   4067: 'Carrier 63 Spacing Fault', class No Acknowledgement, trigger "DB302_HMI_Faults_Carrier63_Faults_2" bit 2
   4068: 'Carrier 63 Duplicate Carrier Number Fault', class No Acknowledgement, trigger "DB302_HMI_Faults_Carrier63_Faults_2" bit 3
   4069: 'Spare_Fault_4069', class No Acknowledgement, trigger "DB302_HMI_Faults_Carrier63_Faults_2" bit 4
   4070: 'Spare_Fault_4070', class No Acknowledgement, trigger "DB302_HMI_Faults_Carrier63_Faults_2" bit 5
   4071: 'Spare_Fault_4071', class No Acknowledgement, trigger "DB302_HMI_Faults_Carrier63_Faults_2" bit 6
   4072: 'Spare_Fault_4072', class No Acknowledgement, trigger "DB302_HMI_Faults_Carrier63_Faults_2" bit 7
   4073: 'Spare_Fault_4073', class No Acknowledgement, trigger "DB302_HMI_Faults_Carrier63_Faults_2" bit 8
   4074: 'Spare_Fault_4074', class No Acknowledgement, trigger "DB302_HMI_Faults_Carrier63_Faults_2" bit 9
   4075: 'Spare_Fault_4075', class No Acknowledgement, trigger "DB302_HMI_Faults_Carrier63_Faults_2" bit 10
   4076: 'Spare_Fault_4076', class No Acknowledgement, trigger "DB302_HMI_Faults_Carrier63_Faults_2" bit 11
   4077: 'Spare_Fault_4077', class No Acknowledgement, trigger "DB302_HMI_Faults_Carrier63_Faults_2" bit 12
   4078: 'Spare_Fault_4078', class No Acknowledgement, trigger "DB302_HMI_Faults_Carrier63_Faults_2" bit 13
   4079: 'Spare_Fault_4079', class No Acknowledgement, trigger "DB302_HMI_Faults_Carrier63_Faults_2" bit 14
   4080: 'Spare_Fault_4080', class No Acknowledgement, trigger "DB302_HMI_Faults_Carrier63_Faults_2" bit 15
   4081: 'Spare_Fault_4081', class No Acknowledgement, trigger "DB302_HMI_Faults_Carrier63_Faults_3" bit 0
   4082: 'Spare_Fault_4082', class No Acknowledgement, trigger "DB302_HMI_Faults_Carrier63_Faults_3" bit 1
   4083: 'Spare_Fault_4083', class No Acknowledgement, trigger "DB302_HMI_Faults_Carrier63_Faults_3" bit 2
   4084: 'Spare_Fault_4084', class No Acknowledgement, trigger "DB302_HMI_Faults_Carrier63_Faults_3" bit 3
   4085: 'Spare_Fault_4085', class No Acknowledgement, trigger "DB302_HMI_Faults_Carrier63_Faults_3" bit 4
   4086: 'Spare_Fault_4086', class No Acknowledgement, trigger "DB302_HMI_Faults_Carrier63_Faults_3" bit 5
   4087: 'Spare_Fault_4087', class No Acknowledgement, trigger "DB302_HMI_Faults_Carrier63_Faults_3" bit 6
   4088: 'Spare_Fault_4088', class No Acknowledgement, trigger "DB302_HMI_Faults_Carrier63_Faults_3" bit 7
   4089: 'Spare_Fault_4089', class No Acknowledgement, trigger "DB302_HMI_Faults_Carrier63_Faults_3" bit 8
   4090: 'Spare_Fault_4090', class No Acknowledgement, trigger "DB302_HMI_Faults_Carrier63_Faults_3" bit 9
   4091: 'Spare_Fault_4091', class No Acknowledgement, trigger "DB302_HMI_Faults_Carrier63_Faults_3" bit 10
   4092: 'Spare_Fault_4092', class No Acknowledgement, trigger "DB302_HMI_Faults_Carrier63_Faults_3" bit 11
   4093: 'Spare_Fault_4093', class No Acknowledgement, trigger "DB302_HMI_Faults_Carrier63_Faults_3" bit 12
   4094: 'Spare_Fault_4094', class No Acknowledgement, trigger "DB302_HMI_Faults_Carrier63_Faults_3" bit 13
   4095: 'Spare_Fault_4095', class No Acknowledgement, trigger "DB302_HMI_Faults_Carrier63_Faults_3" bit 14
   4096: 'Spare_Fault_4096', class No Acknowledgement, trigger "DB302_HMI_Faults_Carrier63_Faults_3" bit 15
   4097: 'Carrier 64 Disconnect Open Power Fault DI11.0', class No Acknowledgement, trigger "DB302_HMI_Faults_Carrier64_Faults_0" bit 0
   4098: 'Carrier 64 Drive Profinet Comm Fault', class No Acknowledgement, trigger "DB302_HMI_Faults_Carrier64_Faults_0" bit 1
   4099: 'Carrier 64 Production Stop Not Reset', class No Acknowledgement, trigger "DB302_HMI_Faults_Carrier64_Faults_0" bit 2
   4100: 'Carrier 64 CB02122 Tripped', class No Acknowledgement, trigger "DB302_HMI_Faults_Carrier64_Faults_0" bit 3
   4101: 'Carrier 64 CB02123 Tripped', class No Acknowledgement, trigger "DB302_HMI_Faults_Carrier64_Faults_0" bit 4
   4102: 'Carrier 64 AUX1 CB Tripped', class No Acknowledgement, trigger "DB302_HMI_Faults_Carrier64_Faults_0" bit 5
   4103: 'Carrier 64 AUX2 CB Tripped', class No Acknowledgement, trigger "DB302_HMI_Faults_Carrier64_Faults_0" bit 6
   4104: 'Carrier 64 PLC Not Communicating', class No Acknowledgement, trigger "DB302_HMI_Faults_Carrier64_Faults_0" bit 7
   4105: 'Carrier 64 Safe Input Card Fault', class No Acknowledgement, trigger "DB302_HMI_Faults_Carrier64_Faults_0" bit 8
   4106: 'Carrier 64 Safe Output Card Fault', class No Acknowledgement, trigger "DB302_HMI_Faults_Carrier64_Faults_0" bit 9
   4107: 'Carrier 64 Standard Input Card Fault', class No Acknowledgement, trigger "DB302_HMI_Faults_Carrier64_Faults_0" bit 10
   4108: 'Carrier 64 Standard Output Card Fault', class No Acknowledgement, trigger "DB302_HMI_Faults_Carrier64_Faults_0" bit 11
   4109: 'Carrier 64 Encoder Position Fault', class No Acknowledgement, trigger "DB302_HMI_Faults_Carrier64_Faults_0" bit 12
   4110: 'Carrier 64 Encoder Internal Error', class No Acknowledgement, trigger "DB302_HMI_Faults_Carrier64_Faults_0" bit 13
   4111: 'Carrier 64 Encoder Comm Fault', class No Acknowledgement, trigger "DB302_HMI_Faults_Carrier64_Faults_0" bit 14
   4112: 'Carrier 64 HMI Comm Fault', class No Acknowledgement, trigger "DB302_HMI_Faults_Carrier64_Faults_0" bit 15
   4113: 'Carrier 64 Crash Detection Fault', class No Acknowledgement, trigger "DB302_HMI_Faults_Carrier64_Faults_1" bit 0
   4114: 'Carrier 64 Carrier Number Invalid', class No Acknowledgement, trigger "DB302_HMI_Faults_Carrier64_Faults_1" bit 1
   4115: 'Carrier 64 Drive: PROFINET configuration error', class No Acknowledgement, trigger "DB302_HMI_Faults_Carrier64_Faults_1" bit 2
   4116: 'Carrier 64 Drive: Error internal communications', class No Acknowledgement, trigger "DB302_HMI_Faults_Carrier64_Faults_1" bit 3
   4117: 'Carrier 64 Drive: Motor overtemperature', class No Acknowledgement, trigger "DB302_HMI_Faults_Carrier64_Faults_1" bit 4
   4118: 'Carrier 64 Drive: Motor overcurrent', class No Acknowledgement, trigger "DB302_HMI_Faults_Carrier64_Faults_1" bit 5
   4119: 'Carrier 64 Drive: Infeed or power unit not ready', class No Acknowledgement, trigger "DB302_HMI_Faults_Carrier64_Faults_1" bit 6
   4120: 'Carrier 64 Drive: Short-circuit/ground fault detected', class No Acknowledgement, trigger "DB302_HMI_Faults_Carrier64_Faults_1" bit 7
   4121: 'Carrier 64 Drive: PROFINET Setpoint timeout', class No Acknowledgement, trigger "DB302_HMI_Faults_Carrier64_Faults_1" bit 8
   4122: 'Carrier 64 Power unit: Overcurrent', class No Acknowledgement, trigger "DB302_HMI_Faults_Carrier64_Faults_1" bit 9
   4123: 'Carrier 64 Power unit: DC link voltage overvoltage', class No Acknowledgement, trigger "DB302_HMI_Faults_Carrier64_Faults_1" bit 10
   4124: 'Carrier 64 Power unit: DC link voltage undervoltage', class No Acknowledgement, trigger "DB302_HMI_Faults_Carrier64_Faults_1" bit 11
   4125: 'Carrier 64 Power unit: Line phase failure in main circuit', class No Acknowledgement, trigger "DB302_HMI_Faults_Carrier64_Faults_1" bit 12
   4126: 'Carrier 64 Power unit: Phase failure motor cable', class No Acknowledgement, trigger "DB302_HMI_Faults_Carrier64_Faults_1" bit 13
   4127: 'Carrier 64 Power unit: Ground fault', class No Acknowledgement, trigger "DB302_HMI_Faults_Carrier64_Faults_1" bit 14
   4128: 'Spare_Fault_4128', class No Acknowledgement, trigger "DB302_HMI_Faults_Carrier64_Faults_1" bit 15
   4129: 'Carrier 64 Motion Off Fault', class No Acknowledgement, trigger "DB302_HMI_Faults_Carrier64_Faults_2" bit 0
   4130: 'Carrier 64 Motion On Fault', class No Acknowledgement, trigger "DB302_HMI_Faults_Carrier64_Faults_2" bit 1
   4131: 'Carrier 64 Spacing Fault', class No Acknowledgement, trigger "DB302_HMI_Faults_Carrier64_Faults_2" bit 2
   4132: 'Carrier 64 Duplicate Carrier Number Fault', class No Acknowledgement, trigger "DB302_HMI_Faults_Carrier64_Faults_2" bit 3
   4133: 'Spare_Fault_4133', class No Acknowledgement, trigger "DB302_HMI_Faults_Carrier64_Faults_2" bit 4
   4134: 'Spare_Fault_4134', class No Acknowledgement, trigger "DB302_HMI_Faults_Carrier64_Faults_2" bit 5
   4135: 'Spare_Fault_4135', class No Acknowledgement, trigger "DB302_HMI_Faults_Carrier64_Faults_2" bit 6
   4136: 'Spare_Fault_4136', class No Acknowledgement, trigger "DB302_HMI_Faults_Carrier64_Faults_2" bit 7
   4137: 'Spare_Fault_4137', class No Acknowledgement, trigger "DB302_HMI_Faults_Carrier64_Faults_2" bit 8
   4138: 'Spare_Fault_4138', class No Acknowledgement, trigger "DB302_HMI_Faults_Carrier64_Faults_2" bit 9
   4139: 'Spare_Fault_4139', class No Acknowledgement, trigger "DB302_HMI_Faults_Carrier64_Faults_2" bit 10
   4140: 'Spare_Fault_4140', class No Acknowledgement, trigger "DB302_HMI_Faults_Carrier64_Faults_2" bit 11
   4141: 'Spare_Fault_4141', class No Acknowledgement, trigger "DB302_HMI_Faults_Carrier64_Faults_2" bit 12
   4142: 'Spare_Fault_4142', class No Acknowledgement, trigger "DB302_HMI_Faults_Carrier64_Faults_2" bit 13
   4143: 'Spare_Fault_4143', class No Acknowledgement, trigger "DB302_HMI_Faults_Carrier64_Faults_2" bit 14
   4144: 'Spare_Fault_4144', class No Acknowledgement, trigger "DB302_HMI_Faults_Carrier64_Faults_2" bit 15
   4145: 'Spare_Fault_4145', class No Acknowledgement, trigger "DB302_HMI_Faults_Carrier64_Faults_3" bit 0
   4146: 'Spare_Fault_4146', class No Acknowledgement, trigger "DB302_HMI_Faults_Carrier64_Faults_3" bit 1
   4147: 'Spare_Fault_4147', class No Acknowledgement, trigger "DB302_HMI_Faults_Carrier64_Faults_3" bit 2
   4148: 'Spare_Fault_4148', class No Acknowledgement, trigger "DB302_HMI_Faults_Carrier64_Faults_3" bit 3
   4149: 'Spare_Fault_4149', class No Acknowledgement, trigger "DB302_HMI_Faults_Carrier64_Faults_3" bit 4
   4150: 'Spare_Fault_4150', class No Acknowledgement, trigger "DB302_HMI_Faults_Carrier64_Faults_3" bit 5
   4151: 'Spare_Fault_4151', class No Acknowledgement, trigger "DB302_HMI_Faults_Carrier64_Faults_3" bit 6
   4152: 'Spare_Fault_4152', class No Acknowledgement, trigger "DB302_HMI_Faults_Carrier64_Faults_3" bit 7
   4153: 'Spare_Fault_4153', class No Acknowledgement, trigger "DB302_HMI_Faults_Carrier64_Faults_3" bit 8
   4154: 'Spare_Fault_4154', class No Acknowledgement, trigger "DB302_HMI_Faults_Carrier64_Faults_3" bit 9
   4155: 'Spare_Fault_4155', class No Acknowledgement, trigger "DB302_HMI_Faults_Carrier64_Faults_3" bit 10
   4156: 'Spare_Fault_4156', class No Acknowledgement, trigger "DB302_HMI_Faults_Carrier64_Faults_3" bit 11
   4157: 'Spare_Fault_4157', class No Acknowledgement, trigger "DB302_HMI_Faults_Carrier64_Faults_3" bit 12
   4158: 'Spare_Fault_4158', class No Acknowledgement, trigger "DB302_HMI_Faults_Carrier64_Faults_3" bit 13
   4159: 'Spare_Fault_4159', class No Acknowledgement, trigger "DB302_HMI_Faults_Carrier64_Faults_3" bit 14
   4160: 'Spare_Fault_4160', class No Acknowledgement, trigger "DB302_HMI_Faults_Carrier64_Faults_3" bit 15
   4161: 'Carrier 65 Disconnect Open Power Fault DI11.0', class No Acknowledgement, trigger "DB302_HMI_Faults_Carrier65_Faults_0" bit 0
   4162: 'Carrier 65 Drive Profinet Comm Fault', class No Acknowledgement, trigger "DB302_HMI_Faults_Carrier65_Faults_0" bit 1
   4163: 'Carrier 65 Production Stop Not Reset', class No Acknowledgement, trigger "DB302_HMI_Faults_Carrier65_Faults_0" bit 2
   4164: 'Carrier 65 CB02122 Tripped', class No Acknowledgement, trigger "DB302_HMI_Faults_Carrier65_Faults_0" bit 3
   4165: 'Carrier 65 CB02123 Tripped', class No Acknowledgement, trigger "DB302_HMI_Faults_Carrier65_Faults_0" bit 4
   4166: 'Carrier 65 AUX1 CB Tripped', class No Acknowledgement, trigger "DB302_HMI_Faults_Carrier65_Faults_0" bit 5
   4167: 'Carrier 65 AUX2 CB Tripped', class No Acknowledgement, trigger "DB302_HMI_Faults_Carrier65_Faults_0" bit 6
   4168: 'Carrier 65 PLC Not Communicating', class No Acknowledgement, trigger "DB302_HMI_Faults_Carrier65_Faults_0" bit 7
   4169: 'Carrier 65 Safe Input Card Fault', class No Acknowledgement, trigger "DB302_HMI_Faults_Carrier65_Faults_0" bit 8
   4170: 'Carrier 65 Safe Output Card Fault', class No Acknowledgement, trigger "DB302_HMI_Faults_Carrier65_Faults_0" bit 9
   4171: 'Carrier 65 Standard Input Card Fault', class No Acknowledgement, trigger "DB302_HMI_Faults_Carrier65_Faults_0" bit 10
   4172: 'Carrier 65 Standard Output Card Fault', class No Acknowledgement, trigger "DB302_HMI_Faults_Carrier65_Faults_0" bit 11
   4173: 'Carrier 65 Encoder Position Fault', class No Acknowledgement, trigger "DB302_HMI_Faults_Carrier65_Faults_0" bit 12
   4174: 'Carrier 65 Encoder Internal Error', class No Acknowledgement, trigger "DB302_HMI_Faults_Carrier65_Faults_0" bit 13
   4175: 'Carrier 65 Encoder Comm Fault', class No Acknowledgement, trigger "DB302_HMI_Faults_Carrier65_Faults_0" bit 14
   4176: 'Carrier 65 HMI Comm Fault', class No Acknowledgement, trigger "DB302_HMI_Faults_Carrier65_Faults_0" bit 15
   4177: 'Carrier 65 Crash Detection Fault', class No Acknowledgement, trigger "DB302_HMI_Faults_Carrier65_Faults_1" bit 0
   4178: 'Carrier 65 Carrier Number Invalid', class No Acknowledgement, trigger "DB302_HMI_Faults_Carrier65_Faults_1" bit 1
   4179: 'Carrier 65 Drive: PROFINET configuration error', class No Acknowledgement, trigger "DB302_HMI_Faults_Carrier65_Faults_1" bit 2
   4180: 'Carrier 65 Drive: Error internal communications', class No Acknowledgement, trigger "DB302_HMI_Faults_Carrier65_Faults_1" bit 3
   4181: 'Carrier 65 Drive: Motor overtemperature', class No Acknowledgement, trigger "DB302_HMI_Faults_Carrier65_Faults_1" bit 4
   4182: 'Carrier 65 Drive: Motor overcurrent', class No Acknowledgement, trigger "DB302_HMI_Faults_Carrier65_Faults_1" bit 5
   4183: 'Carrier 65 Drive: Infeed or power unit not ready', class No Acknowledgement, trigger "DB302_HMI_Faults_Carrier65_Faults_1" bit 6
   4184: 'Carrier 65 Drive: Short-circuit/ground fault detected', class No Acknowledgement, trigger "DB302_HMI_Faults_Carrier65_Faults_1" bit 7
   4185: 'Carrier 65 Drive: PROFINET Setpoint timeout', class No Acknowledgement, trigger "DB302_HMI_Faults_Carrier65_Faults_1" bit 8
   4186: 'Carrier 65 Power unit: Overcurrent', class No Acknowledgement, trigger "DB302_HMI_Faults_Carrier65_Faults_1" bit 9
   4187: 'Carrier 65 Power unit: DC link voltage overvoltage', class No Acknowledgement, trigger "DB302_HMI_Faults_Carrier65_Faults_1" bit 10
   4188: 'Carrier 65 Power unit: DC link voltage undervoltage', class No Acknowledgement, trigger "DB302_HMI_Faults_Carrier65_Faults_1" bit 11
   4189: 'Carrier 65 Power unit: Line phase failure in main circuit', class No Acknowledgement, trigger "DB302_HMI_Faults_Carrier65_Faults_1" bit 12
   4190: 'Carrier 65 Power unit: Phase failure motor cable', class No Acknowledgement, trigger "DB302_HMI_Faults_Carrier65_Faults_1" bit 13
   4191: 'Carrier 65 Power unit: Ground fault', class No Acknowledgement, trigger "DB302_HMI_Faults_Carrier65_Faults_1" bit 14
   4192: 'Spare_Fault_4192', class No Acknowledgement, trigger "DB302_HMI_Faults_Carrier65_Faults_1" bit 15
   4193: 'Carrier 65 Motion Off Fault', class No Acknowledgement, trigger "DB302_HMI_Faults_Carrier65_Faults_2" bit 0
   4194: 'Carrier 65 Motion On Fault', class No Acknowledgement, trigger "DB302_HMI_Faults_Carrier65_Faults_2" bit 1
   4195: 'Carrier 65 Spacing Fault', class No Acknowledgement, trigger "DB302_HMI_Faults_Carrier65_Faults_2" bit 2
   4196: 'Carrier 65 Duplicate Carrier Number Fault', class No Acknowledgement, trigger "DB302_HMI_Faults_Carrier65_Faults_2" bit 3
   4197: 'Spare_Fault_4197', class No Acknowledgement, trigger "DB302_HMI_Faults_Carrier65_Faults_2" bit 4
   4198: 'Spare_Fault_4198', class No Acknowledgement, trigger "DB302_HMI_Faults_Carrier65_Faults_2" bit 5
   4199: 'Spare_Fault_4199', class No Acknowledgement, trigger "DB302_HMI_Faults_Carrier65_Faults_2" bit 6
   4200: 'Spare_Fault_4200', class No Acknowledgement, trigger "DB302_HMI_Faults_Carrier65_Faults_2" bit 7
   4201: 'Spare_Fault_4201', class No Acknowledgement, trigger "DB302_HMI_Faults_Carrier65_Faults_2" bit 8
   4202: 'Spare_Fault_4202', class No Acknowledgement, trigger "DB302_HMI_Faults_Carrier65_Faults_2" bit 9
   4203: 'Spare_Fault_4203', class No Acknowledgement, trigger "DB302_HMI_Faults_Carrier65_Faults_2" bit 10
   4204: 'Spare_Fault_4204', class No Acknowledgement, trigger "DB302_HMI_Faults_Carrier65_Faults_2" bit 11
   4205: 'Spare_Fault_4205', class No Acknowledgement, trigger "DB302_HMI_Faults_Carrier65_Faults_2" bit 12
   4206: 'Spare_Fault_4206', class No Acknowledgement, trigger "DB302_HMI_Faults_Carrier65_Faults_2" bit 13
   4207: 'Spare_Fault_4207', class No Acknowledgement, trigger "DB302_HMI_Faults_Carrier65_Faults_2" bit 14
   4208: 'Spare_Fault_4208', class No Acknowledgement, trigger "DB302_HMI_Faults_Carrier65_Faults_2" bit 15
   4209: 'Spare_Fault_4209', class No Acknowledgement, trigger "DB302_HMI_Faults_Carrier65_Faults_3" bit 0
   4210: 'Spare_Fault_4210', class No Acknowledgement, trigger "DB302_HMI_Faults_Carrier65_Faults_3" bit 1
   4211: 'Spare_Fault_4211', class No Acknowledgement, trigger "DB302_HMI_Faults_Carrier65_Faults_3" bit 2
   4212: 'Spare_Fault_4212', class No Acknowledgement, trigger "DB302_HMI_Faults_Carrier65_Faults_3" bit 3
   4213: 'Spare_Fault_4213', class No Acknowledgement, trigger "DB302_HMI_Faults_Carrier65_Faults_3" bit 4
   4214: 'Spare_Fault_4214', class No Acknowledgement, trigger "DB302_HMI_Faults_Carrier65_Faults_3" bit 5
   4215: 'Spare_Fault_4215', class No Acknowledgement, trigger "DB302_HMI_Faults_Carrier65_Faults_3" bit 6
   4216: 'Spare_Fault_4216', class No Acknowledgement, trigger "DB302_HMI_Faults_Carrier65_Faults_3" bit 7
   4217: 'Spare_Fault_4217', class No Acknowledgement, trigger "DB302_HMI_Faults_Carrier65_Faults_3" bit 8
   4218: 'Spare_Fault_4218', class No Acknowledgement, trigger "DB302_HMI_Faults_Carrier65_Faults_3" bit 9
   4219: 'Spare_Fault_4219', class No Acknowledgement, trigger "DB302_HMI_Faults_Carrier65_Faults_3" bit 10
   4220: 'Spare_Fault_4220', class No Acknowledgement, trigger "DB302_HMI_Faults_Carrier65_Faults_3" bit 11
   4221: 'Spare_Fault_4221', class No Acknowledgement, trigger "DB302_HMI_Faults_Carrier65_Faults_3" bit 12
   4222: 'Spare_Fault_4222', class No Acknowledgement, trigger "DB302_HMI_Faults_Carrier65_Faults_3" bit 13
   4223: 'Spare_Fault_4223', class No Acknowledgement, trigger "DB302_HMI_Faults_Carrier65_Faults_3" bit 14
   4224: 'Spare_Fault_4224', class No Acknowledgement, trigger "DB302_HMI_Faults_Carrier65_Faults_3" bit 15
   4225: 'Carrier 66 Disconnect Open Power Fault DI11.0', class No Acknowledgement, trigger "DB302_HMI_Faults_Carrier66_Faults_0" bit 0
   4226: 'Carrier 66 Drive Profinet Comm Fault', class No Acknowledgement, trigger "DB302_HMI_Faults_Carrier66_Faults_0" bit 1
   4227: 'Carrier 66 Production Stop Not Reset', class No Acknowledgement, trigger "DB302_HMI_Faults_Carrier66_Faults_0" bit 2
   4228: 'Carrier 66 CB02122 Tripped', class No Acknowledgement, trigger "DB302_HMI_Faults_Carrier66_Faults_0" bit 3
   4229: 'Carrier 66 CB02123 Tripped', class No Acknowledgement, trigger "DB302_HMI_Faults_Carrier66_Faults_0" bit 4
   4230: 'Carrier 66 AUX1 CB Tripped', class No Acknowledgement, trigger "DB302_HMI_Faults_Carrier66_Faults_0" bit 5
   4231: 'Carrier 66 AUX2 CB Tripped', class No Acknowledgement, trigger "DB302_HMI_Faults_Carrier66_Faults_0" bit 6
   4232: 'Carrier 66 PLC Not Communicating', class No Acknowledgement, trigger "DB302_HMI_Faults_Carrier66_Faults_0" bit 7
   4233: 'Carrier 66 Safe Input Card Fault', class No Acknowledgement, trigger "DB302_HMI_Faults_Carrier66_Faults_0" bit 8
   4234: 'Carrier 66 Safe Output Card Fault', class No Acknowledgement, trigger "DB302_HMI_Faults_Carrier66_Faults_0" bit 9
   4235: 'Carrier 66 Standard Input Card Fault', class No Acknowledgement, trigger "DB302_HMI_Faults_Carrier66_Faults_0" bit 10
   4236: 'Carrier 66 Standard Output Card Fault', class No Acknowledgement, trigger "DB302_HMI_Faults_Carrier66_Faults_0" bit 11
   4237: 'Carrier 66 Encoder Position Fault', class No Acknowledgement, trigger "DB302_HMI_Faults_Carrier66_Faults_0" bit 12
   4238: 'Carrier 66 Encoder Internal Error', class No Acknowledgement, trigger "DB302_HMI_Faults_Carrier66_Faults_0" bit 13
   4239: 'Carrier 66 Encoder Comm Fault', class No Acknowledgement, trigger "DB302_HMI_Faults_Carrier66_Faults_0" bit 14
   4240: 'Carrier 66 HMI Comm Fault', class No Acknowledgement, trigger "DB302_HMI_Faults_Carrier66_Faults_0" bit 15
   4241: 'Carrier 66 Crash Detection Fault', class No Acknowledgement, trigger "DB302_HMI_Faults_Carrier66_Faults_1" bit 0
   4242: 'Carrier 66 Carrier Number Invalid', class No Acknowledgement, trigger "DB302_HMI_Faults_Carrier66_Faults_1" bit 1
   4243: 'Carrier 66 Drive: PROFINET configuration error', class No Acknowledgement, trigger "DB302_HMI_Faults_Carrier66_Faults_1" bit 2
   4244: 'Carrier 66 Drive: Error internal communications', class No Acknowledgement, trigger "DB302_HMI_Faults_Carrier66_Faults_1" bit 3
   4245: 'Carrier 66 Drive: Motor overtemperature', class No Acknowledgement, trigger "DB302_HMI_Faults_Carrier66_Faults_1" bit 4
   4246: 'Carrier 66 Drive: Motor overcurrent', class No Acknowledgement, trigger "DB302_HMI_Faults_Carrier66_Faults_1" bit 5
   4247: 'Carrier 66 Drive: Infeed or power unit not ready', class No Acknowledgement, trigger "DB302_HMI_Faults_Carrier66_Faults_1" bit 6
   4248: 'Carrier 66 Drive: Short-circuit/ground fault detected', class No Acknowledgement, trigger "DB302_HMI_Faults_Carrier66_Faults_1" bit 7
   4249: 'Carrier 66 Drive: PROFINET Setpoint timeout', class No Acknowledgement, trigger "DB302_HMI_Faults_Carrier66_Faults_1" bit 8
   4250: 'Carrier 66 Power unit: Overcurrent', class No Acknowledgement, trigger "DB302_HMI_Faults_Carrier66_Faults_1" bit 9
   4251: 'Carrier 66 Power unit: DC link voltage overvoltage', class No Acknowledgement, trigger "DB302_HMI_Faults_Carrier66_Faults_1" bit 10
   4252: 'Carrier 66 Power unit: DC link voltage undervoltage', class No Acknowledgement, trigger "DB302_HMI_Faults_Carrier66_Faults_1" bit 11
   4253: 'Carrier 66 Power unit: Line phase failure in main circuit', class No Acknowledgement, trigger "DB302_HMI_Faults_Carrier66_Faults_1" bit 12
   4254: 'Carrier 66 Power unit: Phase failure motor cable', class No Acknowledgement, trigger "DB302_HMI_Faults_Carrier66_Faults_1" bit 13
   4255: 'Carrier 66 Power unit: Ground fault', class No Acknowledgement, trigger "DB302_HMI_Faults_Carrier66_Faults_1" bit 14
   4256: 'Spare_Fault_4256', class No Acknowledgement, trigger "DB302_HMI_Faults_Carrier66_Faults_1" bit 15
   4257: 'Carrier 66 Motion Off Fault', class No Acknowledgement, trigger "DB302_HMI_Faults_Carrier66_Faults_2" bit 0
   4258: 'Carrier 66 Motion On Fault', class No Acknowledgement, trigger "DB302_HMI_Faults_Carrier66_Faults_2" bit 1
   4259: 'Carrier 66 Spacing Fault', class No Acknowledgement, trigger "DB302_HMI_Faults_Carrier66_Faults_2" bit 2
   4260: 'Carrier 66 Duplicate Carrier Number Fault', class No Acknowledgement, trigger "DB302_HMI_Faults_Carrier66_Faults_2" bit 3
   4261: 'Spare_Fault_4261', class No Acknowledgement, trigger "DB302_HMI_Faults_Carrier66_Faults_2" bit 4
   4262: 'Spare_Fault_4262', class No Acknowledgement, trigger "DB302_HMI_Faults_Carrier66_Faults_2" bit 5
   4263: 'Spare_Fault_4263', class No Acknowledgement, trigger "DB302_HMI_Faults_Carrier66_Faults_2" bit 6
   4264: 'Spare_Fault_4264', class No Acknowledgement, trigger "DB302_HMI_Faults_Carrier66_Faults_2" bit 7
   4265: 'Spare_Fault_4265', class No Acknowledgement, trigger "DB302_HMI_Faults_Carrier66_Faults_2" bit 8
   4266: 'Spare_Fault_4266', class No Acknowledgement, trigger "DB302_HMI_Faults_Carrier66_Faults_2" bit 9
   4267: 'Spare_Fault_4267', class No Acknowledgement, trigger "DB302_HMI_Faults_Carrier66_Faults_2" bit 10
   4268: 'Spare_Fault_4268', class No Acknowledgement, trigger "DB302_HMI_Faults_Carrier66_Faults_2" bit 11
   4269: 'Spare_Fault_4269', class No Acknowledgement, trigger "DB302_HMI_Faults_Carrier66_Faults_2" bit 12
   4270: 'Spare_Fault_4270', class No Acknowledgement, trigger "DB302_HMI_Faults_Carrier66_Faults_2" bit 13
   4271: 'Spare_Fault_4271', class No Acknowledgement, trigger "DB302_HMI_Faults_Carrier66_Faults_2" bit 14
   4272: 'Spare_Fault_4272', class No Acknowledgement, trigger "DB302_HMI_Faults_Carrier66_Faults_2" bit 15
   4273: 'Spare_Fault_4273', class No Acknowledgement, trigger "DB302_HMI_Faults_Carrier66_Faults_3" bit 0
   4274: 'Spare_Fault_4274', class No Acknowledgement, trigger "DB302_HMI_Faults_Carrier66_Faults_3" bit 1
   4275: 'Spare_Fault_4275', class No Acknowledgement, trigger "DB302_HMI_Faults_Carrier66_Faults_3" bit 2
   4276: 'Spare_Fault_4276', class No Acknowledgement, trigger "DB302_HMI_Faults_Carrier66_Faults_3" bit 3
   4277: 'Spare_Fault_4277', class No Acknowledgement, trigger "DB302_HMI_Faults_Carrier66_Faults_3" bit 4
   4278: 'Spare_Fault_4278', class No Acknowledgement, trigger "DB302_HMI_Faults_Carrier66_Faults_3" bit 5
   4279: 'Spare_Fault_4279', class No Acknowledgement, trigger "DB302_HMI_Faults_Carrier66_Faults_3" bit 6
   4280: 'Spare_Fault_4280', class No Acknowledgement, trigger "DB302_HMI_Faults_Carrier66_Faults_3" bit 7
   4281: 'Spare_Fault_4281', class No Acknowledgement, trigger "DB302_HMI_Faults_Carrier66_Faults_3" bit 8
   4282: 'Spare_Fault_4282', class No Acknowledgement, trigger "DB302_HMI_Faults_Carrier66_Faults_3" bit 9
   4283: 'Spare_Fault_4283', class No Acknowledgement, trigger "DB302_HMI_Faults_Carrier66_Faults_3" bit 10
   4284: 'Spare_Fault_4284', class No Acknowledgement, trigger "DB302_HMI_Faults_Carrier66_Faults_3" bit 11
   4285: 'Spare_Fault_4285', class No Acknowledgement, trigger "DB302_HMI_Faults_Carrier66_Faults_3" bit 12
   4286: 'Spare_Fault_4286', class No Acknowledgement, trigger "DB302_HMI_Faults_Carrier66_Faults_3" bit 13
   4287: 'Spare_Fault_4287', class No Acknowledgement, trigger "DB302_HMI_Faults_Carrier66_Faults_3" bit 14
   4288: 'Spare_Fault_4288', class No Acknowledgement, trigger "DB302_HMI_Faults_Carrier66_Faults_3" bit 15
   4289: 'Carrier 67 Disconnect Open Power Fault DI11.0', class No Acknowledgement, trigger "DB302_HMI_Faults_Carrier67_Faults_0" bit 0
   4290: 'Carrier 67 Drive Profinet Comm Fault', class No Acknowledgement, trigger "DB302_HMI_Faults_Carrier67_Faults_0" bit 1
   4291: 'Carrier 67 Production Stop Not Reset', class No Acknowledgement, trigger "DB302_HMI_Faults_Carrier67_Faults_0" bit 2
   4292: 'Carrier 67 CB02122 Tripped', class No Acknowledgement, trigger "DB302_HMI_Faults_Carrier67_Faults_0" bit 3
   4293: 'Carrier 67 CB02123 Tripped', class No Acknowledgement, trigger "DB302_HMI_Faults_Carrier67_Faults_0" bit 4
   4294: 'Carrier 67 AUX1 CB Tripped', class No Acknowledgement, trigger "DB302_HMI_Faults_Carrier67_Faults_0" bit 5
   4295: 'Carrier 67 AUX2 CB Tripped', class No Acknowledgement, trigger "DB302_HMI_Faults_Carrier67_Faults_0" bit 6
   4296: 'Carrier 67 PLC Not Communicating', class No Acknowledgement, trigger "DB302_HMI_Faults_Carrier67_Faults_0" bit 7
   4297: 'Carrier 67 Safe Input Card Fault', class No Acknowledgement, trigger "DB302_HMI_Faults_Carrier67_Faults_0" bit 8
   4298: 'Carrier 67 Safe Output Card Fault', class No Acknowledgement, trigger "DB302_HMI_Faults_Carrier67_Faults_0" bit 9
   4299: 'Carrier 67 Standard Input Card Fault', class No Acknowledgement, trigger "DB302_HMI_Faults_Carrier67_Faults_0" bit 10
   4300: 'Carrier 67 Standard Output Card Fault', class No Acknowledgement, trigger "DB302_HMI_Faults_Carrier67_Faults_0" bit 11
   4301: 'Carrier 67 Encoder Position Fault', class No Acknowledgement, trigger "DB302_HMI_Faults_Carrier67_Faults_0" bit 12
   4302: 'Carrier 67 Encoder Internal Error', class No Acknowledgement, trigger "DB302_HMI_Faults_Carrier67_Faults_0" bit 13
   4303: 'Carrier 67 Encoder Comm Fault', class No Acknowledgement, trigger "DB302_HMI_Faults_Carrier67_Faults_0" bit 14
   4304: 'Carrier 67 HMI Comm Fault', class No Acknowledgement, trigger "DB302_HMI_Faults_Carrier67_Faults_0" bit 15
   4305: 'Carrier 67 Crash Detection Fault', class No Acknowledgement, trigger "DB302_HMI_Faults_Carrier67_Faults_1" bit 0
   4306: 'Carrier 67 Carrier Number Invalid', class No Acknowledgement, trigger "DB302_HMI_Faults_Carrier67_Faults_1" bit 1
   4307: 'Carrier 67 Drive: PROFINET configuration error', class No Acknowledgement, trigger "DB302_HMI_Faults_Carrier67_Faults_1" bit 2
   4308: 'Carrier 67 Drive: Error internal communications', class No Acknowledgement, trigger "DB302_HMI_Faults_Carrier67_Faults_1" bit 3
   4309: 'Carrier 67 Drive: Motor overtemperature', class No Acknowledgement, trigger "DB302_HMI_Faults_Carrier67_Faults_1" bit 4
   4310: 'Carrier 67 Drive: Motor overcurrent', class No Acknowledgement, trigger "DB302_HMI_Faults_Carrier67_Faults_1" bit 5
   4311: 'Carrier 67 Drive: Infeed or power unit not ready', class No Acknowledgement, trigger "DB302_HMI_Faults_Carrier67_Faults_1" bit 6
   4312: 'Carrier 67 Drive: Short-circuit/ground fault detected', class No Acknowledgement, trigger "DB302_HMI_Faults_Carrier67_Faults_1" bit 7
   4313: 'Carrier 67 Drive: PROFINET Setpoint timeout', class No Acknowledgement, trigger "DB302_HMI_Faults_Carrier67_Faults_1" bit 8
   4314: 'Carrier 67 Power unit: Overcurrent', class No Acknowledgement, trigger "DB302_HMI_Faults_Carrier67_Faults_1" bit 9
   4315: 'Carrier 67 Power unit: DC link voltage overvoltage', class No Acknowledgement, trigger "DB302_HMI_Faults_Carrier67_Faults_1" bit 10
   4316: 'Carrier 67 Power unit: DC link voltage undervoltage', class No Acknowledgement, trigger "DB302_HMI_Faults_Carrier67_Faults_1" bit 11
   4317: 'Carrier 67 Power unit: Line phase failure in main circuit', class No Acknowledgement, trigger "DB302_HMI_Faults_Carrier67_Faults_1" bit 12
   4318: 'Carrier 67 Power unit: Phase failure motor cable', class No Acknowledgement, trigger "DB302_HMI_Faults_Carrier67_Faults_1" bit 13
   4319: 'Carrier 67 Power unit: Ground fault', class No Acknowledgement, trigger "DB302_HMI_Faults_Carrier67_Faults_1" bit 14
   4320: 'Spare_Fault_4320', class No Acknowledgement, trigger "DB302_HMI_Faults_Carrier67_Faults_1" bit 15
   4321: 'Carrier 67 Motion Off Fault', class No Acknowledgement, trigger "DB302_HMI_Faults_Carrier67_Faults_2" bit 0
   4322: 'Carrier 67 Motion On Fault', class No Acknowledgement, trigger "DB302_HMI_Faults_Carrier67_Faults_2" bit 1
   4323: 'Carrier 67 Spacing Fault', class No Acknowledgement, trigger "DB302_HMI_Faults_Carrier67_Faults_2" bit 2
   4324: 'Carrier 67 Duplicate Carrier Number Fault', class No Acknowledgement, trigger "DB302_HMI_Faults_Carrier67_Faults_2" bit 3
   4325: 'Spare_Fault_4325', class No Acknowledgement, trigger "DB302_HMI_Faults_Carrier67_Faults_2" bit 4
   4326: 'Spare_Fault_4326', class No Acknowledgement, trigger "DB302_HMI_Faults_Carrier67_Faults_2" bit 5
   4327: 'Spare_Fault_4327', class No Acknowledgement, trigger "DB302_HMI_Faults_Carrier67_Faults_2" bit 6
   4328: 'Spare_Fault_4328', class No Acknowledgement, trigger "DB302_HMI_Faults_Carrier67_Faults_2" bit 7
   4329: 'Spare_Fault_4329', class No Acknowledgement, trigger "DB302_HMI_Faults_Carrier67_Faults_2" bit 8
   4330: 'Spare_Fault_4330', class No Acknowledgement, trigger "DB302_HMI_Faults_Carrier67_Faults_2" bit 9
   4331: 'Spare_Fault_4331', class No Acknowledgement, trigger "DB302_HMI_Faults_Carrier67_Faults_2" bit 10
   4332: 'Spare_Fault_4332', class No Acknowledgement, trigger "DB302_HMI_Faults_Carrier67_Faults_2" bit 11
   4333: 'Spare_Fault_4333', class No Acknowledgement, trigger "DB302_HMI_Faults_Carrier67_Faults_2" bit 12
   4334: 'Spare_Fault_4334', class No Acknowledgement, trigger "DB302_HMI_Faults_Carrier67_Faults_2" bit 13
   4335: 'Spare_Fault_4335', class No Acknowledgement, trigger "DB302_HMI_Faults_Carrier67_Faults_2" bit 14
   4336: 'Spare_Fault_4336', class No Acknowledgement, trigger "DB302_HMI_Faults_Carrier67_Faults_2" bit 15
   4337: 'Spare_Fault_4337', class No Acknowledgement, trigger "DB302_HMI_Faults_Carrier67_Faults_3" bit 0
   4338: 'Spare_Fault_4338', class No Acknowledgement, trigger "DB302_HMI_Faults_Carrier67_Faults_3" bit 1
   4339: 'Spare_Fault_4339', class No Acknowledgement, trigger "DB302_HMI_Faults_Carrier67_Faults_3" bit 2
   4340: 'Spare_Fault_4340', class No Acknowledgement, trigger "DB302_HMI_Faults_Carrier67_Faults_3" bit 3
   4341: 'Spare_Fault_4341', class No Acknowledgement, trigger "DB302_HMI_Faults_Carrier67_Faults_3" bit 4
   4342: 'Spare_Fault_4342', class No Acknowledgement, trigger "DB302_HMI_Faults_Carrier67_Faults_3" bit 5
   4343: 'Spare_Fault_4343', class No Acknowledgement, trigger "DB302_HMI_Faults_Carrier67_Faults_3" bit 6
   4344: 'Spare_Fault_4344', class No Acknowledgement, trigger "DB302_HMI_Faults_Carrier67_Faults_3" bit 7
   4345: 'Spare_Fault_4345', class No Acknowledgement, trigger "DB302_HMI_Faults_Carrier67_Faults_3" bit 8
   4346: 'Spare_Fault_4346', class No Acknowledgement, trigger "DB302_HMI_Faults_Carrier67_Faults_3" bit 9
   4347: 'Spare_Fault_4347', class No Acknowledgement, trigger "DB302_HMI_Faults_Carrier67_Faults_3" bit 10
   4348: 'Spare_Fault_4348', class No Acknowledgement, trigger "DB302_HMI_Faults_Carrier67_Faults_3" bit 11
   4349: 'Spare_Fault_4349', class No Acknowledgement, trigger "DB302_HMI_Faults_Carrier67_Faults_3" bit 12
   4350: 'Spare_Fault_4350', class No Acknowledgement, trigger "DB302_HMI_Faults_Carrier67_Faults_3" bit 13
   4351: 'Spare_Fault_4351', class No Acknowledgement, trigger "DB302_HMI_Faults_Carrier67_Faults_3" bit 14
   4352: 'Spare_Fault_4352', class No Acknowledgement, trigger "DB302_HMI_Faults_Carrier67_Faults_3" bit 15
   4353: 'Carrier 68 Disconnect Open Power Fault DI11.0', class No Acknowledgement, trigger "DB302_HMI_Faults_Carrier68_Faults_0" bit 0
   4354: 'Carrier 68 Drive Profinet Comm Fault', class No Acknowledgement, trigger "DB302_HMI_Faults_Carrier68_Faults_0" bit 1
   4355: 'Carrier 68 Production Stop Not Reset', class No Acknowledgement, trigger "DB302_HMI_Faults_Carrier68_Faults_0" bit 2
   4356: 'Carrier 68 CB02122 Tripped', class No Acknowledgement, trigger "DB302_HMI_Faults_Carrier68_Faults_0" bit 3
   4357: 'Carrier 68 CB02123 Tripped', class No Acknowledgement, trigger "DB302_HMI_Faults_Carrier68_Faults_0" bit 4
   4358: 'Carrier 68 AUX1 CB Tripped', class No Acknowledgement, trigger "DB302_HMI_Faults_Carrier68_Faults_0" bit 5
   4359: 'Carrier 68 AUX2 CB Tripped', class No Acknowledgement, trigger "DB302_HMI_Faults_Carrier68_Faults_0" bit 6
   4360: 'Carrier 68 PLC Not Communicating', class No Acknowledgement, trigger "DB302_HMI_Faults_Carrier68_Faults_0" bit 7
   4361: 'Carrier 68 Safe Input Card Fault', class No Acknowledgement, trigger "DB302_HMI_Faults_Carrier68_Faults_0" bit 8
   4362: 'Carrier 68 Safe Output Card Fault', class No Acknowledgement, trigger "DB302_HMI_Faults_Carrier68_Faults_0" bit 9
   4363: 'Carrier 68 Standard Input Card Fault', class No Acknowledgement, trigger "DB302_HMI_Faults_Carrier68_Faults_0" bit 10
   4364: 'Carrier 68 Standard Output Card Fault', class No Acknowledgement, trigger "DB302_HMI_Faults_Carrier68_Faults_0" bit 11
   4365: 'Carrier 68 Encoder Position Fault', class No Acknowledgement, trigger "DB302_HMI_Faults_Carrier68_Faults_0" bit 12
   4366: 'Carrier 68 Encoder Internal Error', class No Acknowledgement, trigger "DB302_HMI_Faults_Carrier68_Faults_0" bit 13
   4367: 'Carrier 68 Encoder Comm Fault', class No Acknowledgement, trigger "DB302_HMI_Faults_Carrier68_Faults_0" bit 14
   4368: 'Carrier 68 HMI Comm Fault', class No Acknowledgement, trigger "DB302_HMI_Faults_Carrier68_Faults_0" bit 15
   4369: 'Carrier 68 Crash Detection Fault', class No Acknowledgement, trigger "DB302_HMI_Faults_Carrier68_Faults_1" bit 0
   4370: 'Carrier 68 Carrier Number Invalid', class No Acknowledgement, trigger "DB302_HMI_Faults_Carrier68_Faults_1" bit 1
   4371: 'Carrier 68 Drive: PROFINET configuration error', class No Acknowledgement, trigger "DB302_HMI_Faults_Carrier68_Faults_1" bit 2
   4372: 'Carrier 68 Drive: Error internal communications', class No Acknowledgement, trigger "DB302_HMI_Faults_Carrier68_Faults_1" bit 3
   4373: 'Carrier 68 Drive: Motor overtemperature', class No Acknowledgement, trigger "DB302_HMI_Faults_Carrier68_Faults_1" bit 4
   4374: 'Carrier 68 Drive: Motor overcurrent', class No Acknowledgement, trigger "DB302_HMI_Faults_Carrier68_Faults_1" bit 5
   4375: 'Carrier 68 Drive: Infeed or power unit not ready', class No Acknowledgement, trigger "DB302_HMI_Faults_Carrier68_Faults_1" bit 6
   4376: 'Carrier 68 Drive: Short-circuit/ground fault detected', class No Acknowledgement, trigger "DB302_HMI_Faults_Carrier68_Faults_1" bit 7
   4377: 'Carrier 68 Drive: PROFINET Setpoint timeout', class No Acknowledgement, trigger "DB302_HMI_Faults_Carrier68_Faults_1" bit 8
   4378: 'Carrier 68 Power unit: Overcurrent', class No Acknowledgement, trigger "DB302_HMI_Faults_Carrier68_Faults_1" bit 9
   4379: 'Carrier 68 Power unit: DC link voltage overvoltage', class No Acknowledgement, trigger "DB302_HMI_Faults_Carrier68_Faults_1" bit 10
   4380: 'Carrier 68 Power unit: DC link voltage undervoltage', class No Acknowledgement, trigger "DB302_HMI_Faults_Carrier68_Faults_1" bit 11
   4381: 'Carrier 68 Power unit: Line phase failure in main circuit', class No Acknowledgement, trigger "DB302_HMI_Faults_Carrier68_Faults_1" bit 12
   4382: 'Carrier 68 Power unit: Phase failure motor cable', class No Acknowledgement, trigger "DB302_HMI_Faults_Carrier68_Faults_1" bit 13
   4383: 'Carrier 68 Power unit: Ground fault', class No Acknowledgement, trigger "DB302_HMI_Faults_Carrier68_Faults_1" bit 14
   4384: 'Spare_Fault_4384', class No Acknowledgement, trigger "DB302_HMI_Faults_Carrier68_Faults_1" bit 15
   4385: 'Carrier 68 Motion Off Fault', class No Acknowledgement, trigger "DB302_HMI_Faults_Carrier68_Faults_2" bit 0
   4386: 'Carrier 68 Motion On Fault', class No Acknowledgement, trigger "DB302_HMI_Faults_Carrier68_Faults_2" bit 1
   4387: 'Carrier 68 Spacing Fault', class No Acknowledgement, trigger "DB302_HMI_Faults_Carrier68_Faults_2" bit 2
   4388: 'Carrier 68 Duplicate Carrier Number Fault', class No Acknowledgement, trigger "DB302_HMI_Faults_Carrier68_Faults_2" bit 3
   4389: 'Spare_Fault_4389', class No Acknowledgement, trigger "DB302_HMI_Faults_Carrier68_Faults_2" bit 4
   4390: 'Spare_Fault_4390', class No Acknowledgement, trigger "DB302_HMI_Faults_Carrier68_Faults_2" bit 5
   4391: 'Spare_Fault_4391', class No Acknowledgement, trigger "DB302_HMI_Faults_Carrier68_Faults_2" bit 6
   4392: 'Spare_Fault_4392', class No Acknowledgement, trigger "DB302_HMI_Faults_Carrier68_Faults_2" bit 7
   4393: 'Spare_Fault_4393', class No Acknowledgement, trigger "DB302_HMI_Faults_Carrier68_Faults_2" bit 8
   4394: 'Spare_Fault_4394', class No Acknowledgement, trigger "DB302_HMI_Faults_Carrier68_Faults_2" bit 9
   4395: 'Spare_Fault_4395', class No Acknowledgement, trigger "DB302_HMI_Faults_Carrier68_Faults_2" bit 10
   4396: 'Spare_Fault_4396', class No Acknowledgement, trigger "DB302_HMI_Faults_Carrier68_Faults_2" bit 11
   4397: 'Spare_Fault_4397', class No Acknowledgement, trigger "DB302_HMI_Faults_Carrier68_Faults_2" bit 12
   4398: 'Spare_Fault_4398', class No Acknowledgement, trigger "DB302_HMI_Faults_Carrier68_Faults_2" bit 13
   4399: 'Spare_Fault_4399', class No Acknowledgement, trigger "DB302_HMI_Faults_Carrier68_Faults_2" bit 14
   4400: 'Spare_Fault_4400', class No Acknowledgement, trigger "DB302_HMI_Faults_Carrier68_Faults_2" bit 15
   4401: 'Spare_Fault_4401', class No Acknowledgement, trigger "DB302_HMI_Faults_Carrier68_Faults_3" bit 0
   4402: 'Spare_Fault_4402', class No Acknowledgement, trigger "DB302_HMI_Faults_Carrier68_Faults_3" bit 1
   4403: 'Spare_Fault_4403', class No Acknowledgement, trigger "DB302_HMI_Faults_Carrier68_Faults_3" bit 2
   4404: 'Spare_Fault_4404', class No Acknowledgement, trigger "DB302_HMI_Faults_Carrier68_Faults_3" bit 3
   4405: 'Spare_Fault_4405', class No Acknowledgement, trigger "DB302_HMI_Faults_Carrier68_Faults_3" bit 4
   4406: 'Spare_Fault_4406', class No Acknowledgement, trigger "DB302_HMI_Faults_Carrier68_Faults_3" bit 5
   4407: 'Spare_Fault_4407', class No Acknowledgement, trigger "DB302_HMI_Faults_Carrier68_Faults_3" bit 6
   4408: 'Spare_Fault_4408', class No Acknowledgement, trigger "DB302_HMI_Faults_Carrier68_Faults_3" bit 7
   4409: 'Spare_Fault_4409', class No Acknowledgement, trigger "DB302_HMI_Faults_Carrier68_Faults_3" bit 8
   4410: 'Spare_Fault_4410', class No Acknowledgement, trigger "DB302_HMI_Faults_Carrier68_Faults_3" bit 9
   4411: 'Spare_Fault_4411', class No Acknowledgement, trigger "DB302_HMI_Faults_Carrier68_Faults_3" bit 10
   4412: 'Spare_Fault_4412', class No Acknowledgement, trigger "DB302_HMI_Faults_Carrier68_Faults_3" bit 11
   4413: 'Spare_Fault_4413', class No Acknowledgement, trigger "DB302_HMI_Faults_Carrier68_Faults_3" bit 12
   4414: 'Spare_Fault_4414', class No Acknowledgement, trigger "DB302_HMI_Faults_Carrier68_Faults_3" bit 13
   4415: 'Spare_Fault_4415', class No Acknowledgement, trigger "DB302_HMI_Faults_Carrier68_Faults_3" bit 14
   4416: 'Spare_Fault_4416', class No Acknowledgement, trigger "DB302_HMI_Faults_Carrier68_Faults_3" bit 15
   4417: 'Carrier 69 Disconnect Open Power Fault DI11.0', class No Acknowledgement, trigger "DB302_HMI_Faults_Carrier69_Faults_0" bit 0
   4418: 'Carrier 69 Drive Profinet Comm Fault', class No Acknowledgement, trigger "DB302_HMI_Faults_Carrier69_Faults_0" bit 1
   4419: 'Carrier 69 Production Stop Not Reset', class No Acknowledgement, trigger "DB302_HMI_Faults_Carrier69_Faults_0" bit 2
   4420: 'Carrier 69 CB02122 Tripped', class No Acknowledgement, trigger "DB302_HMI_Faults_Carrier69_Faults_0" bit 3
   4421: 'Carrier 69 CB02123 Tripped', class No Acknowledgement, trigger "DB302_HMI_Faults_Carrier69_Faults_0" bit 4
   4422: 'Carrier 69 AUX1 CB Tripped', class No Acknowledgement, trigger "DB302_HMI_Faults_Carrier69_Faults_0" bit 5
   4423: 'Carrier 69 AUX2 CB Tripped', class No Acknowledgement, trigger "DB302_HMI_Faults_Carrier69_Faults_0" bit 6
   4424: 'Carrier 69 PLC Not Communicating', class No Acknowledgement, trigger "DB302_HMI_Faults_Carrier69_Faults_0" bit 7
   4425: 'Carrier 69 Safe Input Card Fault', class No Acknowledgement, trigger "DB302_HMI_Faults_Carrier69_Faults_0" bit 8
   4426: 'Carrier 69 Safe Output Card Fault', class No Acknowledgement, trigger "DB302_HMI_Faults_Carrier69_Faults_0" bit 9
   4427: 'Carrier 69 Standard Input Card Fault', class No Acknowledgement, trigger "DB302_HMI_Faults_Carrier69_Faults_0" bit 10
   4428: 'Carrier 69 Standard Output Card Fault', class No Acknowledgement, trigger "DB302_HMI_Faults_Carrier69_Faults_0" bit 11
   4429: 'Carrier 69 Encoder Position Fault', class No Acknowledgement, trigger "DB302_HMI_Faults_Carrier69_Faults_0" bit 12
   4430: 'Carrier 69 Encoder Internal Error', class No Acknowledgement, trigger "DB302_HMI_Faults_Carrier69_Faults_0" bit 13
   4431: 'Carrier 69 Encoder Comm Fault', class No Acknowledgement, trigger "DB302_HMI_Faults_Carrier69_Faults_0" bit 14
   4432: 'Carrier 69 HMI Comm Fault', class No Acknowledgement, trigger "DB302_HMI_Faults_Carrier69_Faults_0" bit 15
   4433: 'Carrier 69 Crash Detection Fault', class No Acknowledgement, trigger "DB302_HMI_Faults_Carrier69_Faults_1" bit 0
   4434: 'Carrier 69 Carrier Number Invalid', class No Acknowledgement, trigger "DB302_HMI_Faults_Carrier69_Faults_1" bit 1
   4435: 'Carrier 69 Drive: PROFINET configuration error', class No Acknowledgement, trigger "DB302_HMI_Faults_Carrier69_Faults_1" bit 2
   4436: 'Carrier 69 Drive: Error internal communications', class No Acknowledgement, trigger "DB302_HMI_Faults_Carrier69_Faults_1" bit 3
   4437: 'Carrier 69 Drive: Motor overtemperature', class No Acknowledgement, trigger "DB302_HMI_Faults_Carrier69_Faults_1" bit 4
   4438: 'Carrier 69 Drive: Motor overcurrent', class No Acknowledgement, trigger "DB302_HMI_Faults_Carrier69_Faults_1" bit 5
   4439: 'Carrier 69 Drive: Infeed or power unit not ready', class No Acknowledgement, trigger "DB302_HMI_Faults_Carrier69_Faults_1" bit 6
   4440: 'Carrier 69 Drive: Short-circuit/ground fault detected', class No Acknowledgement, trigger "DB302_HMI_Faults_Carrier69_Faults_1" bit 7
   4441: 'Carrier 69 Drive: PROFINET Setpoint timeout', class No Acknowledgement, trigger "DB302_HMI_Faults_Carrier69_Faults_1" bit 8
   4442: 'Carrier 69 Power unit: Overcurrent', class No Acknowledgement, trigger "DB302_HMI_Faults_Carrier69_Faults_1" bit 9
   4443: 'Carrier 69 Power unit: DC link voltage overvoltage', class No Acknowledgement, trigger "DB302_HMI_Faults_Carrier69_Faults_1" bit 10
   4444: 'Carrier 69 Power unit: DC link voltage undervoltage', class No Acknowledgement, trigger "DB302_HMI_Faults_Carrier69_Faults_1" bit 11
   4445: 'Carrier 69 Power unit: Line phase failure in main circuit', class No Acknowledgement, trigger "DB302_HMI_Faults_Carrier69_Faults_1" bit 12
   4446: 'Carrier 69 Power unit: Phase failure motor cable', class No Acknowledgement, trigger "DB302_HMI_Faults_Carrier69_Faults_1" bit 13
   4447: 'Carrier 69 Power unit: Ground fault', class No Acknowledgement, trigger "DB302_HMI_Faults_Carrier69_Faults_1" bit 14
   4448: 'Spare_Fault_4448', class No Acknowledgement, trigger "DB302_HMI_Faults_Carrier69_Faults_1" bit 15
   4449: 'Carrier 69 Motion Off Fault', class No Acknowledgement, trigger "DB302_HMI_Faults_Carrier69_Faults_2" bit 0
   4450: 'Carrier 69 Motion On Fault', class No Acknowledgement, trigger "DB302_HMI_Faults_Carrier69_Faults_2" bit 1
   4451: 'Carrier 69 Spacing Fault', class No Acknowledgement, trigger "DB302_HMI_Faults_Carrier69_Faults_2" bit 2
   4452: 'Carrier 69 Duplicate Carrier Number Fault', class No Acknowledgement, trigger "DB302_HMI_Faults_Carrier69_Faults_2" bit 3
   4453: 'Spare_Fault_4453', class No Acknowledgement, trigger "DB302_HMI_Faults_Carrier69_Faults_2" bit 4
   4454: 'Spare_Fault_4454', class No Acknowledgement, trigger "DB302_HMI_Faults_Carrier69_Faults_2" bit 5
   4455: 'Spare_Fault_4455', class No Acknowledgement, trigger "DB302_HMI_Faults_Carrier69_Faults_2" bit 6
   4456: 'Spare_Fault_4456', class No Acknowledgement, trigger "DB302_HMI_Faults_Carrier69_Faults_2" bit 7
   4457: 'Spare_Fault_4457', class No Acknowledgement, trigger "DB302_HMI_Faults_Carrier69_Faults_2" bit 8
   4458: 'Spare_Fault_4458', class No Acknowledgement, trigger "DB302_HMI_Faults_Carrier69_Faults_2" bit 9
   4459: 'Spare_Fault_4459', class No Acknowledgement, trigger "DB302_HMI_Faults_Carrier69_Faults_2" bit 10
   4460: 'Spare_Fault_4460', class No Acknowledgement, trigger "DB302_HMI_Faults_Carrier69_Faults_2" bit 11
   4461: 'Spare_Fault_4461', class No Acknowledgement, trigger "DB302_HMI_Faults_Carrier69_Faults_2" bit 12
   4462: 'Spare_Fault_4462', class No Acknowledgement, trigger "DB302_HMI_Faults_Carrier69_Faults_2" bit 13
   4463: 'Spare_Fault_4463', class No Acknowledgement, trigger "DB302_HMI_Faults_Carrier69_Faults_2" bit 14
   4464: 'Spare_Fault_4464', class No Acknowledgement, trigger "DB302_HMI_Faults_Carrier69_Faults_2" bit 15
   4465: 'Spare_Fault_4465', class No Acknowledgement, trigger "DB302_HMI_Faults_Carrier69_Faults_3" bit 0
   4466: 'Spare_Fault_4466', class No Acknowledgement, trigger "DB302_HMI_Faults_Carrier69_Faults_3" bit 1
   4467: 'Spare_Fault_4467', class No Acknowledgement, trigger "DB302_HMI_Faults_Carrier69_Faults_3" bit 2
   4468: 'Spare_Fault_4468', class No Acknowledgement, trigger "DB302_HMI_Faults_Carrier69_Faults_3" bit 3
   4469: 'Spare_Fault_4469', class No Acknowledgement, trigger "DB302_HMI_Faults_Carrier69_Faults_3" bit 4
   4470: 'Spare_Fault_4470', class No Acknowledgement, trigger "DB302_HMI_Faults_Carrier69_Faults_3" bit 5
   4471: 'Spare_Fault_4471', class No Acknowledgement, trigger "DB302_HMI_Faults_Carrier69_Faults_3" bit 6
   4472: 'Spare_Fault_4472', class No Acknowledgement, trigger "DB302_HMI_Faults_Carrier69_Faults_3" bit 7
   4473: 'Spare_Fault_4473', class No Acknowledgement, trigger "DB302_HMI_Faults_Carrier69_Faults_3" bit 8
   4474: 'Spare_Fault_4474', class No Acknowledgement, trigger "DB302_HMI_Faults_Carrier69_Faults_3" bit 9
   4475: 'Spare_Fault_4475', class No Acknowledgement, trigger "DB302_HMI_Faults_Carrier69_Faults_3" bit 10
   4476: 'Spare_Fault_4476', class No Acknowledgement, trigger "DB302_HMI_Faults_Carrier69_Faults_3" bit 11
   4477: 'Spare_Fault_4477', class No Acknowledgement, trigger "DB302_HMI_Faults_Carrier69_Faults_3" bit 12
   4478: 'Spare_Fault_4478', class No Acknowledgement, trigger "DB302_HMI_Faults_Carrier69_Faults_3" bit 13
   4479: 'Spare_Fault_4479', class No Acknowledgement, trigger "DB302_HMI_Faults_Carrier69_Faults_3" bit 14
   4480: 'Spare_Fault_4480', class No Acknowledgement, trigger "DB302_HMI_Faults_Carrier69_Faults_3" bit 15
   4481: 'Carrier 70 Disconnect Open Power Fault DI11.0', class No Acknowledgement, trigger "DB302_HMI_Faults_Carrier70_Faults_0" bit 0
   4482: 'Carrier 70 Drive Profinet Comm Fault', class No Acknowledgement, trigger "DB302_HMI_Faults_Carrier70_Faults_0" bit 1
   4483: 'Carrier 70 Production Stop Not Reset', class No Acknowledgement, trigger "DB302_HMI_Faults_Carrier70_Faults_0" bit 2
   4484: 'Carrier 70 CB02122 Tripped', class No Acknowledgement, trigger "DB302_HMI_Faults_Carrier70_Faults_0" bit 3
   4485: 'Carrier 70 CB02123 Tripped', class No Acknowledgement, trigger "DB302_HMI_Faults_Carrier70_Faults_0" bit 4
   4486: 'Carrier 70 AUX1 CB Tripped', class No Acknowledgement, trigger "DB302_HMI_Faults_Carrier70_Faults_0" bit 5
   4487: 'Carrier 70 AUX2 CB Tripped', class No Acknowledgement, trigger "DB302_HMI_Faults_Carrier70_Faults_0" bit 6
   4488: 'Carrier 70 PLC Not Communicating', class No Acknowledgement, trigger "DB302_HMI_Faults_Carrier70_Faults_0" bit 7
   4489: 'Carrier 70 Safe Input Card Fault', class No Acknowledgement, trigger "DB302_HMI_Faults_Carrier70_Faults_0" bit 8
   4490: 'Carrier 70 Safe Output Card Fault', class No Acknowledgement, trigger "DB302_HMI_Faults_Carrier70_Faults_0" bit 9